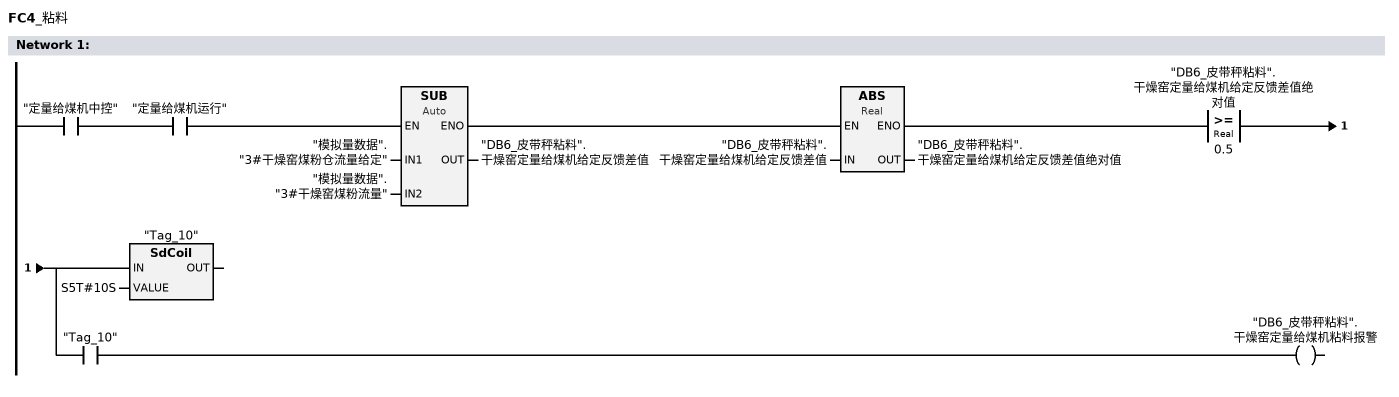
   // no SCL statement known for SdCoil: written as a call
   #_w1 := "定量给煤机中控" AND "定量给煤机运行";
   IF #_w1 THEN
       "DB6_皮带秤粘料".干燥窑定量给煤机给定反馈差值 := "模拟量数据"."3#干燥窑煤粉仓流量给定" - "模拟量数据"."3#干燥窑煤粉流量";
       "DB6_皮带秤粘料".干燥窑定量给煤机给定反馈差值绝对值 := ABS("DB6_皮带秤粘料".干燥窑定量给煤机给定反馈差值);
   END_IF;
   #_w2 := #_w1 AND ("DB6_皮带秤粘料".干燥窑定量给煤机给定反馈差值绝对值 >= 0.5);
   SdCoil(in := #_w2, value := S5T#10S, operand := "Tag_10");
   "DB6_皮带秤粘料".干燥窑定量给煤机粘料报警 := #_w2 AND "Tag_10";
END_REGION
END_FUNCTION

FUNCTION "澳泰温度巡检仪" : Void   // FC5, LAD
{ S7_Optimized_Access := 'FALSE' }
VERSION : 0.1
BEGIN

REGION Network 1
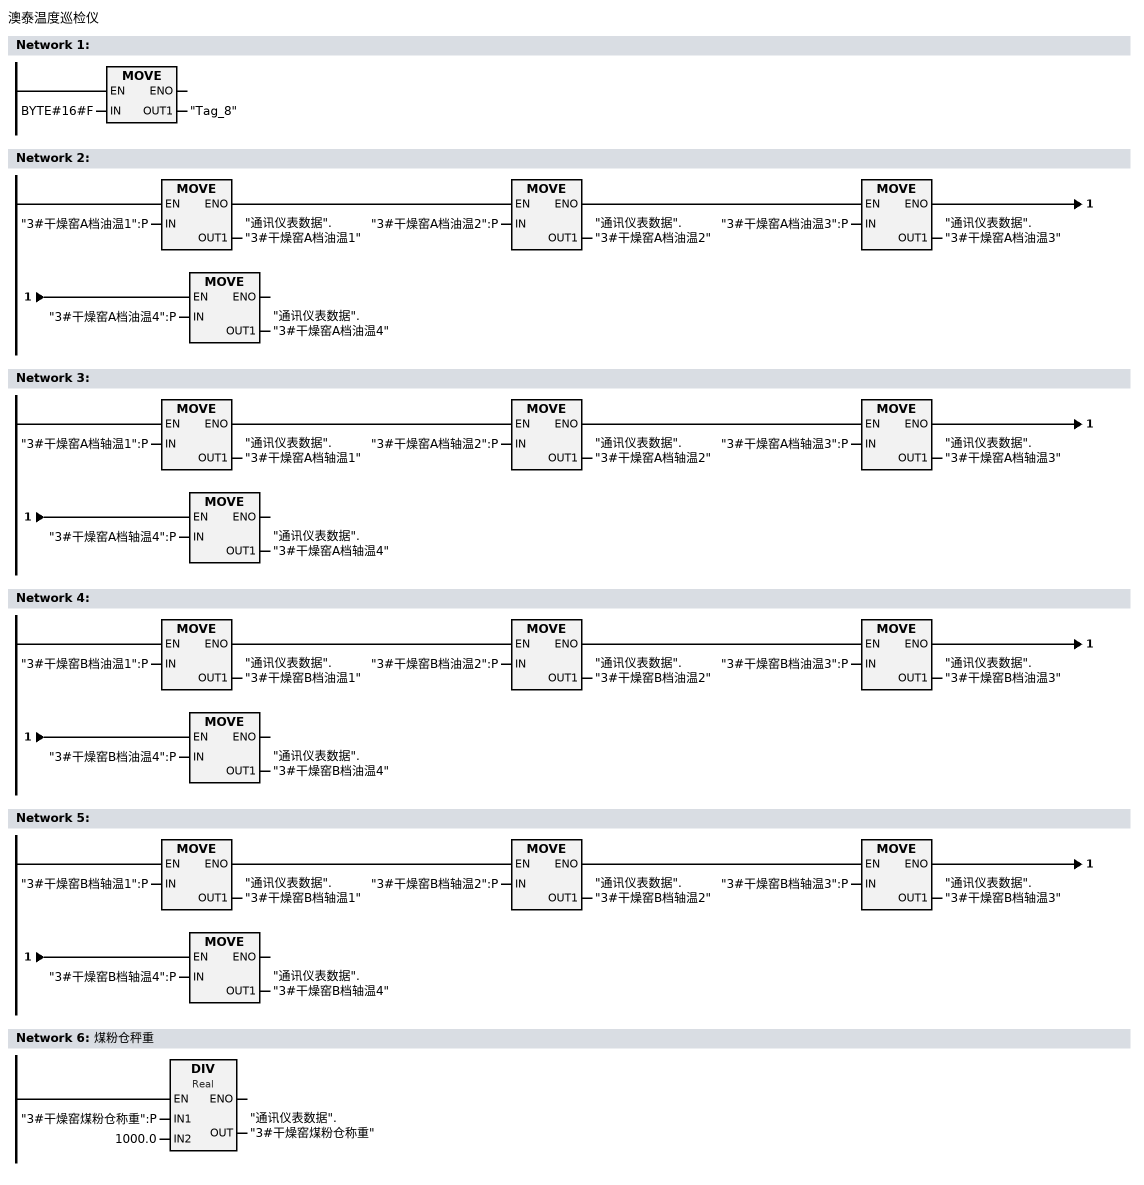
   RUNG wire#powerrail
      { S7_GenerateENO := "TRUE" } Move(in := BYTE#16#F, out1 => "Tag_8")
   END_RUNG
   // the same network as SCL:
   "Tag_8" := BYTE#16#F;
END_REGION

REGION Network 2
   RUNG wire#powerrail
      { S7_GenerateENO := "TRUE" } Move(in := "3#干燥窑A档油温1":P, out1 => "通讯仪表数据"."3#干燥窑A档油温1")
      { S7_GenerateENO := "TRUE" } Move(in := "3#干燥窑A档油温2":P, out1 => "通讯仪表数据"."3#干燥窑A档油温2")
      { S7_GenerateENO := "TRUE" } Move(in := "3#干燥窑A档油温3":P, out1 => "通讯仪表数据"."3#干燥窑A档油温3")
      { S7_GenerateENO := "TRUE" } Move(in := "3#干燥窑A档油温4":P, out1 => "通讯仪表数据"."3#干燥窑A档油温4")
   END_RUNG
   // the same network as SCL:
   // ENO of a box is taken as its EN; it also drops when the box reports an error
   "通讯仪表数据"."3#干燥窑A档油温1" := "3#干燥窑A档油温1":P;
   "通讯仪表数据"."3#干燥窑A档油温2" := "3#干燥窑A档油温2":P;
   "通讯仪表数据"."3#干燥窑A档油温3" := "3#干燥窑A档油温3":P;
   "通讯仪表数据"."3#干燥窑A档油温4" := "3#干燥窑A档油温4":P;
END_REGION

REGION Network 3
   RUNG wire#powerrail
      { S7_GenerateENO := "TRUE" } Move(in := "3#干燥窑A档轴温1":P, out1 => "通讯仪表数据"."3#干燥窑A档轴温1")
      { S7_GenerateENO := "TRUE" } Move(in := "3#干燥窑A档轴温2":P, out1 => "通讯仪表数据"."3#干燥窑A档轴温2")
      { S7_GenerateENO := "TRUE" } Move(in := "3#干燥窑A档轴温3":P, out1 => "通讯仪表数据"."3#干燥窑A档轴温3")
      { S7_GenerateENO := "TRUE" } Move(in := "3#干燥窑A档轴温4":P, out1 => "通讯仪表数据"."3#干燥窑A档轴温4")
   END_RUNG
   // the same network as SCL:
   // ENO of a box is taken as its EN; it also drops when the box reports an error
   "通讯仪表数据"."3#干燥窑A档轴温1" := "3#干燥窑A档轴温1":P;
   "通讯仪表数据"."3#干燥窑A档轴温2" := "3#干燥窑A档轴温2":P;
   "通讯仪表数据"."3#干燥窑A档轴温3" := "3#干燥窑A档轴温3":P;
   "通讯仪表数据"."3#干燥窑A档轴温4" := "3#干燥窑A档轴温4":P;
END_REGION

REGION Network 4
   RUNG wire#powerrail
      { S7_GenerateENO := "TRUE" } Move(in := "3#干燥窑B档油温1":P, out1 => "通讯仪表数据"."3#干燥窑B档油温1")
      { S7_GenerateENO := "TRUE" } Move(in := "3#干燥窑B档油温2":P, out1 => "通讯仪表数据"."3#干燥窑B档油温2")
      { S7_GenerateENO := "TRUE" } Move(in := "3#干燥窑B档油温3":P, out1 => "通讯仪表数据"."3#干燥窑B档油温3")
      { S7_GenerateENO := "TRUE" } Move(in := "3#干燥窑B档油温4":P, out1 => "通讯仪表数据"."3#干燥窑B档油温4")
   END_RUNG
   // the same network as SCL:
   // ENO of a box is taken as its EN; it also drops when the box reports an error
   "通讯仪表数据"."3#干燥窑B档油温1" := "3#干燥窑B档油温1":P;
   "通讯仪表数据"."3#干燥窑B档油温2" := "3#干燥窑B档油温2":P;
   "通讯仪表数据"."3#干燥窑B档油温3" := "3#干燥窑B档油温3":P;
   "通讯仪表数据"."3#干燥窑B档油温4" := "3#干燥窑B档油温4":P;
END_REGION

REGION Network 5
   RUNG wire#powerrail
      { S7_GenerateENO := "TRUE" } Move(in := "3#干燥窑B档轴温1":P, out1 => "通讯仪表数据"."3#干燥窑B档轴温1")
      { S7_GenerateENO := "TRUE" } Move(in := "3#干燥窑B档轴温2":P, out1 => "通讯仪表数据"."3#干燥窑B档轴温2")
      { S7_GenerateENO := "TRUE" } Move(in := "3#干燥窑B档轴温3":P, out1 => "通讯仪表数据"."3#干燥窑B档轴温3")
      { S7_GenerateENO := "TRUE" } Move(in := "3#干燥窑B档轴温4":P, out1 => "通讯仪表数据"."3#干燥窑B档轴温4")
   END_RUNG
   // the same network as SCL:
   // ENO of a box is taken as its EN; it also drops when the box reports an error
   "通讯仪表数据"."3#干燥窑B档轴温1" := "3#干燥窑B档轴温1":P;
   "通讯仪表数据"."3#干燥窑B档轴温2" := "3#干燥窑B档轴温2":P;
   "通讯仪表数据"."3#干燥窑B档轴温3" := "3#干燥窑B档轴温3":P;
   "通讯仪表数据"."3#干燥窑B档轴温4" := "3#干燥窑B档轴温4":P;
END_REGION

REGION Network 6: 煤粉仓秤重
   RUNG wire#powerrail
      { S7_Templates := "SrcType := Real" } Div(in1 := "3#干燥窑煤粉仓称重":P, in2 := 1000.0, out => "通讯仪表数据"."3#干燥窑煤粉仓称重")
   END_RUNG
   // the same network as SCL:
   "通讯仪表数据"."3#干燥窑煤粉仓称重" := "3#干燥窑煤粉仓称重":P / 1000.0;
END_REGION
END_FUNCTION

FUNCTION "3#4#干燥窑皮带联锁信号" : Void   // FC16, LAD
{ S7_Optimized_Access := 'FALSE' }
VERSION : 0.1
BEGIN

REGION Network 1
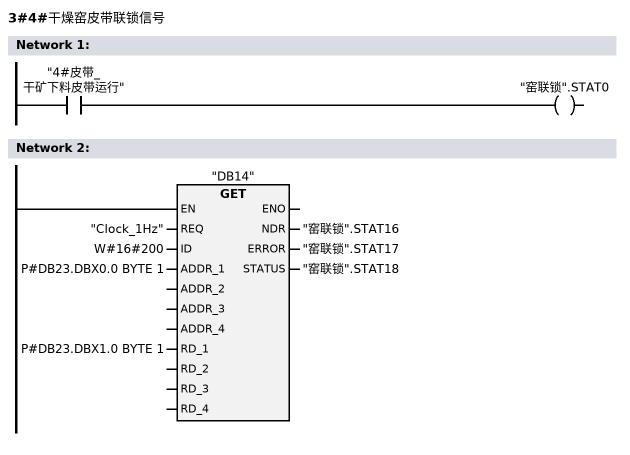
   RUNG wire#powerrail
      Contact( "4#皮带_干矿下料皮带运行" )
      Coil( "窑联锁".STAT0 )
   END_RUNG
   // the same network as SCL:
   "窑联锁".STAT0 := "4#皮带_干矿下料皮带运行";
END_REGION

REGION Network 2
   "DB14"(REQ := "Clock_1Hz",   // GET
          ID := W#16#200,
          ADDR_1 := P#DB23.DBX0.0 BYTE 1,
          RD_1 := P#DB23.DBX1.0 BYTE 1,
          NDR => "窑联锁".STAT16,
          ERROR => "窑联锁".STAT17,
          STATUS => "窑联锁".STAT18);
END_REGION
END_FUNCTION

FUNCTION "模拟量转换" : Void   // FC21, LAD
{ S7_Optimized_Access := 'FALSE' }
VERSION : 0.1
BEGIN

REGION Network 1
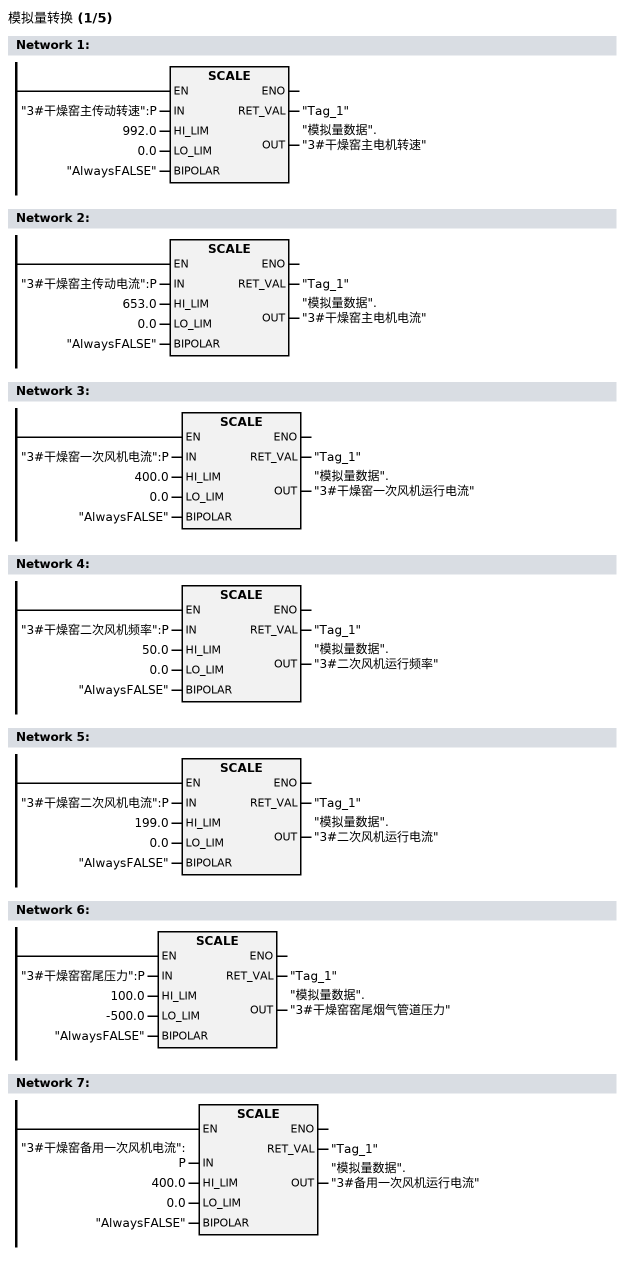
   "Tag_1" := SCALE(IN := "3#干燥窑主传动转速":P,
                    HI_LIM := 992.0,
                    LO_LIM := 0.0,
                    BIPOLAR := "AlwaysFALSE",
                    OUT => "模拟量数据"."3#干燥窑主电机转速");
END_REGION

REGION Network 2
   "Tag_1" := SCALE(IN := "3#干燥窑主传动电流":P,
                    HI_LIM := 653.0,
                    LO_LIM := 0.0,
                    BIPOLAR := "AlwaysFALSE",
                    OUT => "模拟量数据"."3#干燥窑主电机电流");
END_REGION

REGION Network 3
   "Tag_1" := SCALE(IN := "3#干燥窑一次风机电流":P,
                    HI_LIM := 400.0,
                    LO_LIM := 0.0,
                    BIPOLAR := "AlwaysFALSE",
                    OUT => "模拟量数据"."3#干燥窑一次风机运行电流");
END_REGION

REGION Network 4
   "Tag_1" := SCALE(IN := "3#干燥窑二次风机频率":P,
                    HI_LIM := 50.0,
                    LO_LIM := 0.0,
                    BIPOLAR := "AlwaysFALSE",
                    OUT => "模拟量数据"."3#二次风机运行频率");
END_REGION

REGION Network 5
   "Tag_1" := SCALE(IN := "3#干燥窑二次风机电流":P,
                    HI_LIM := 199.0,
                    LO_LIM := 0.0,
                    BIPOLAR := "AlwaysFALSE",
                    OUT => "模拟量数据"."3#二次风机运行电流");
END_REGION

REGION Network 6
   "Tag_1" := SCALE(IN := "3#干燥窑窑尾压力":P,
                    HI_LIM := 100.0,
                    LO_LIM := -500.0,
                    BIPOLAR := "AlwaysFALSE",
                    OUT => "模拟量数据"."3#干燥窑窑尾烟气管道压力");
END_REGION

REGION Network 7
   "Tag_1" := SCALE(IN := "3#干燥窑备用一次风机电流":P,
                    HI_LIM := 400.0,
                    LO_LIM := 0.0,
                    BIPOLAR := "AlwaysFALSE",
                    OUT => "模拟量数据"."3#备用一次风机运行电流");
END_REGION

REGION Network 8
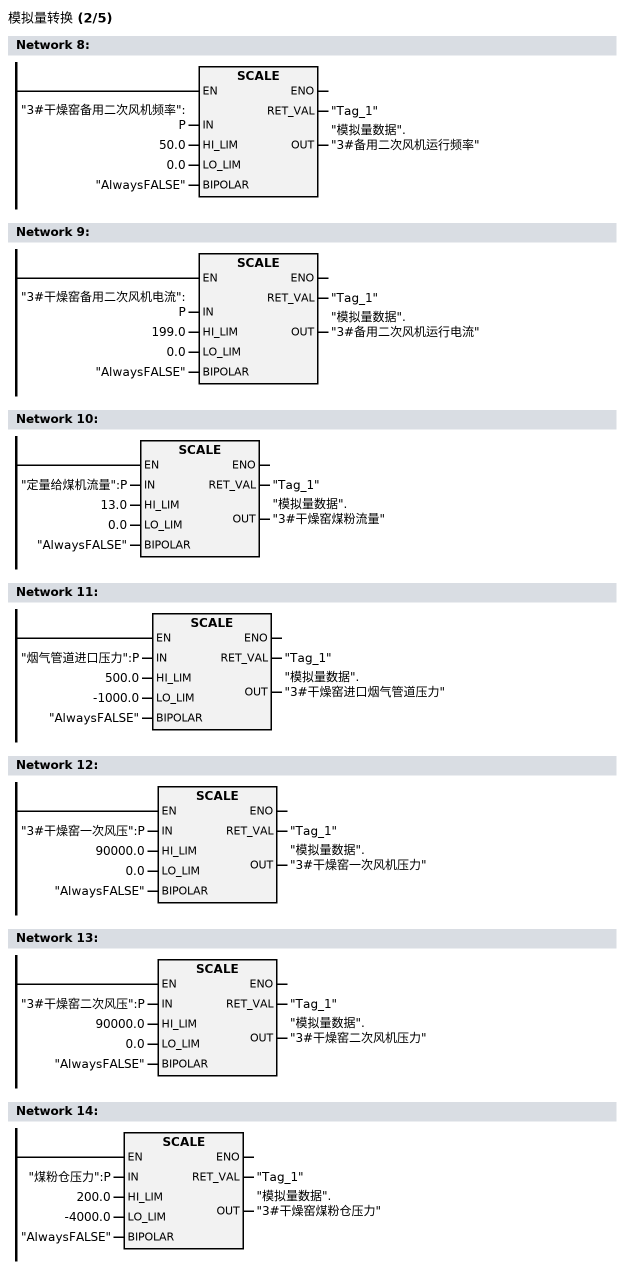
   "Tag_1" := SCALE(IN := "3#干燥窑备用二次风机频率":P,
                    HI_LIM := 50.0,
                    LO_LIM := 0.0,
                    BIPOLAR := "AlwaysFALSE",
                    OUT => "模拟量数据"."3#备用二次风机运行频率");
END_REGION

REGION Network 9
   "Tag_1" := SCALE(IN := "3#干燥窑备用二次风机电流":P,
                    HI_LIM := 199.0,
                    LO_LIM := 0.0,
                    BIPOLAR := "AlwaysFALSE",
                    OUT => "模拟量数据"."3#备用二次风机运行电流");
END_REGION

REGION Network 10
   "Tag_1" := SCALE(IN := "定量给煤机流量":P,
                    HI_LIM := 13.0,
                    LO_LIM := 0.0,
                    BIPOLAR := "AlwaysFALSE",
                    OUT => "模拟量数据"."3#干燥窑煤粉流量");
END_REGION

REGION Network 11
   "Tag_1" := SCALE(IN := "烟气管道进口压力":P,
                    HI_LIM := 500.0,
                    LO_LIM := -1000.0,
                    BIPOLAR := "AlwaysFALSE",
                    OUT => "模拟量数据"."3#干燥窑进口烟气管道压力");
END_REGION

REGION Network 12
   "Tag_1" := SCALE(IN := "3#干燥窑一次风压":P,
                    HI_LIM := 90000.0,
                    LO_LIM := 0.0,
                    BIPOLAR := "AlwaysFALSE",
                    OUT => "模拟量数据"."3#干燥窑一次风机压力");
END_REGION

REGION Network 13
   "Tag_1" := SCALE(IN := "3#干燥窑二次风压":P,
                    HI_LIM := 90000.0,
                    LO_LIM := 0.0,
                    BIPOLAR := "AlwaysFALSE",
                    OUT => "模拟量数据"."3#干燥窑二次风机压力");
END_REGION

REGION Network 14
   "Tag_1" := SCALE(IN := "煤粉仓压力":P,
                    HI_LIM := 200.0,
                    LO_LIM := -4000.0,
                    BIPOLAR := "AlwaysFALSE",
                    OUT => "模拟量数据"."3#干燥窑煤粉仓压力");
END_REGION

REGION Network 15
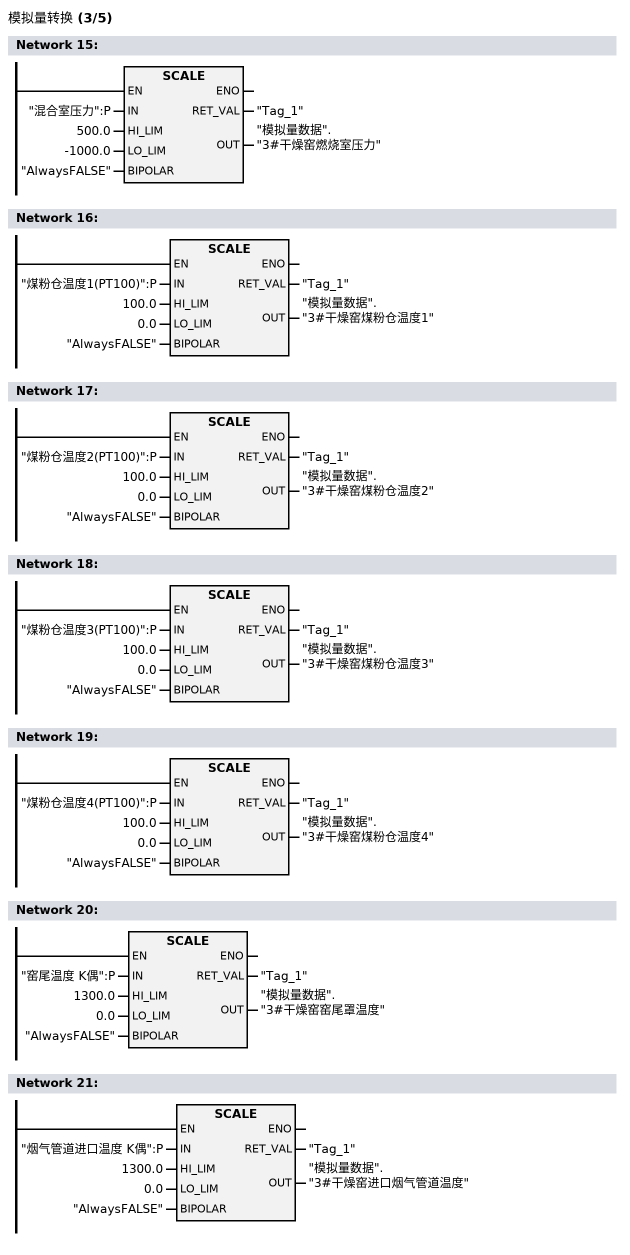
   "Tag_1" := SCALE(IN := "混合室压力":P,
                    HI_LIM := 500.0,
                    LO_LIM := -1000.0,
                    BIPOLAR := "AlwaysFALSE",
                    OUT => "模拟量数据"."3#干燥窑燃烧室压力");
END_REGION

REGION Network 16
   "Tag_1" := SCALE(IN := "煤粉仓温度1(PT100)":P,
                    HI_LIM := 100.0,
                    LO_LIM := 0.0,
                    BIPOLAR := "AlwaysFALSE",
                    OUT => "模拟量数据"."3#干燥窑煤粉仓温度1");
END_REGION

REGION Network 17
   "Tag_1" := SCALE(IN := "煤粉仓温度2(PT100)":P,
                    HI_LIM := 100.0,
                    LO_LIM := 0.0,
                    BIPOLAR := "AlwaysFALSE",
                    OUT => "模拟量数据"."3#干燥窑煤粉仓温度2");
END_REGION

REGION Network 18
   "Tag_1" := SCALE(IN := "煤粉仓温度3(PT100)":P,
                    HI_LIM := 100.0,
                    LO_LIM := 0.0,
                    BIPOLAR := "AlwaysFALSE",
                    OUT => "模拟量数据"."3#干燥窑煤粉仓温度3");
END_REGION

REGION Network 19
   "Tag_1" := SCALE(IN := "煤粉仓温度4(PT100)":P,
                    HI_LIM := 100.0,
                    LO_LIM := 0.0,
                    BIPOLAR := "AlwaysFALSE",
                    OUT => "模拟量数据"."3#干燥窑煤粉仓温度4");
END_REGION

REGION Network 20
   "Tag_1" := SCALE(IN := "窑尾温度 K偶":P,
                    HI_LIM := 1300.0,
                    LO_LIM := 0.0,
                    BIPOLAR := "AlwaysFALSE",
                    OUT => "模拟量数据"."3#干燥窑窑尾罩温度");
END_REGION

REGION Network 21
   "Tag_1" := SCALE(IN := "烟气管道进口温度 K偶":P,
                    HI_LIM := 1300.0,
                    LO_LIM := 0.0,
                    BIPOLAR := "AlwaysFALSE",
                    OUT => "模拟量数据"."3#干燥窑进口烟气管道温度");
END_REGION

REGION Network 22
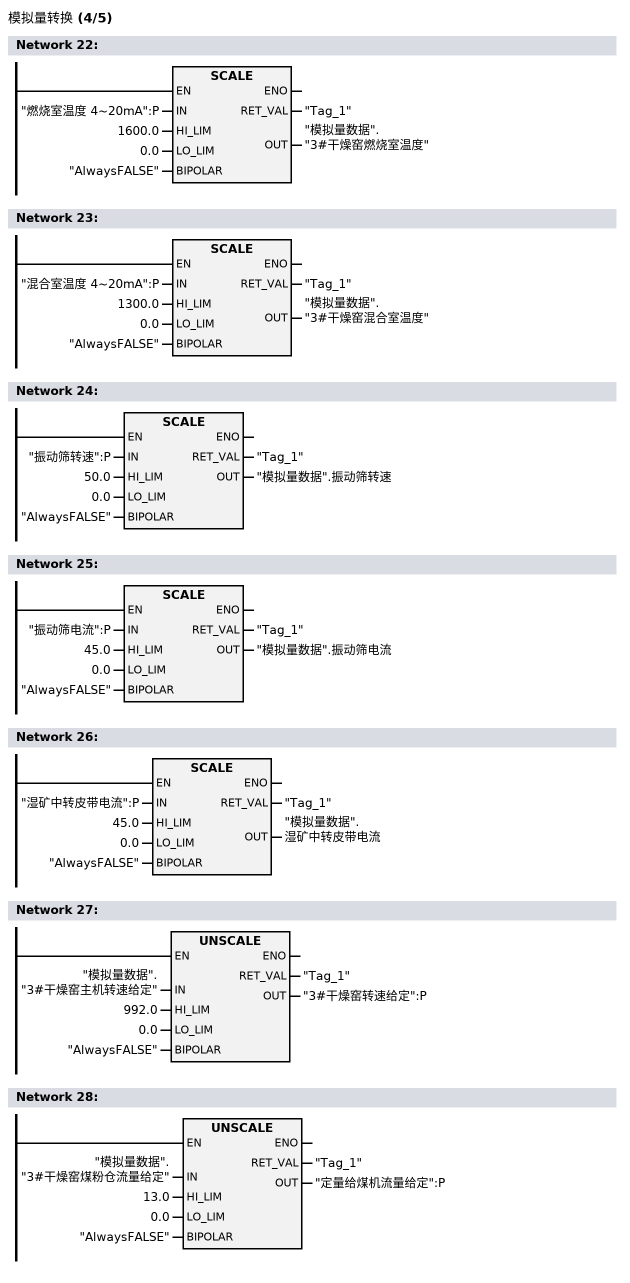
   "Tag_1" := SCALE(IN := "燃烧室温度 4~20mA":P,
                    HI_LIM := 1600.0,
                    LO_LIM := 0.0,
                    BIPOLAR := "AlwaysFALSE",
                    OUT => "模拟量数据"."3#干燥窑燃烧室温度");
END_REGION

REGION Network 23
   "Tag_1" := SCALE(IN := "混合室温度 4~20mA":P,
                    HI_LIM := 1300.0,
                    LO_LIM := 0.0,
                    BIPOLAR := "AlwaysFALSE",
                    OUT => "模拟量数据"."3#干燥窑混合室温度");
END_REGION

REGION Network 24
   "Tag_1" := SCALE(IN := "振动筛转速":P,
                    HI_LIM := 50.0,
                    LO_LIM := 0.0,
                    BIPOLAR := "AlwaysFALSE",
                    OUT => "模拟量数据".振动筛转速);
END_REGION

REGION Network 25
   "Tag_1" := SCALE(IN := "振动筛电流":P,
                    HI_LIM := 45.0,
                    LO_LIM := 0.0,
                    BIPOLAR := "AlwaysFALSE",
                    OUT => "模拟量数据".振动筛电流);
END_REGION

REGION Network 26
   "Tag_1" := SCALE(IN := "湿矿中转皮带电流":P,
                    HI_LIM := 45.0,
                    LO_LIM := 0.0,
                    BIPOLAR := "AlwaysFALSE",
                    OUT => "模拟量数据".湿矿中转皮带电流);
END_REGION

REGION Network 27
   "Tag_1" := UNSCALE(IN := "模拟量数据"."3#干燥窑主机转速给定",
                      HI_LIM := 992.0,
                      LO_LIM := 0.0,
                      BIPOLAR := "AlwaysFALSE",
                      OUT => "3#干燥窑转速给定":P);
END_REGION

REGION Network 28
   "Tag_1" := UNSCALE(IN := "模拟量数据"."3#干燥窑煤粉仓流量给定",
                      HI_LIM := 13.0,
                      LO_LIM := 0.0,
                      BIPOLAR := "AlwaysFALSE",
                      OUT => "定量给煤机流量给定":P);
END_REGION

REGION Network 29
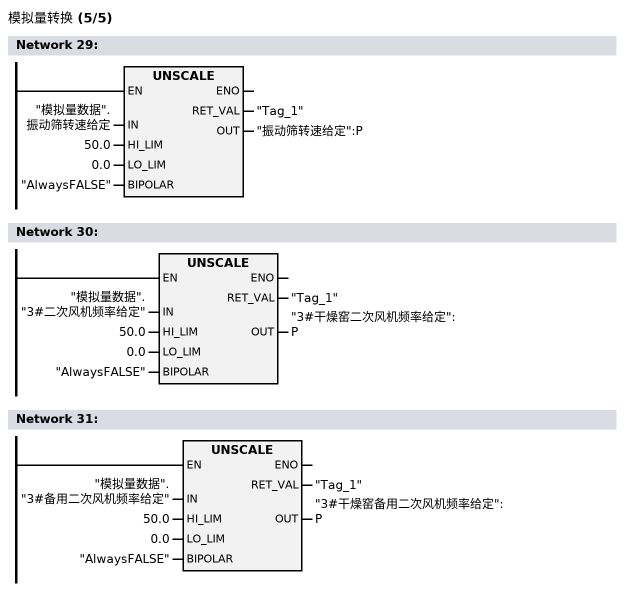
   "Tag_1" := UNSCALE(IN := "模拟量数据".振动筛转速给定,
                      HI_LIM := 50.0,
                      LO_LIM := 0.0,
                      BIPOLAR := "AlwaysFALSE",
                      OUT => "振动筛转速给定":P);
END_REGION

REGION Network 30
   "Tag_1" := UNSCALE(IN := "模拟量数据"."3#二次风机频率给定",
                      HI_LIM := 50.0,
                      LO_LIM := 0.0,
                      BIPOLAR := "AlwaysFALSE",
                      OUT => "3#干燥窑二次风机频率给定":P);
END_REGION

REGION Network 31
   "Tag_1" := UNSCALE(IN := "模拟量数据"."3#备用二次风机频率给定",
                      HI_LIM := 50.0,
                      LO_LIM := 0.0,
                      BIPOLAR := "AlwaysFALSE",
                      OUT => "3#干燥窑备用二次风机频率给定":P);
END_REGION
END_FUNCTION

FUNCTION "皮带机" : Void   // FC22, LAD
{ S7_Optimized_Access := 'FALSE' }
VERSION : 0.1
BEGIN

REGION Network 1
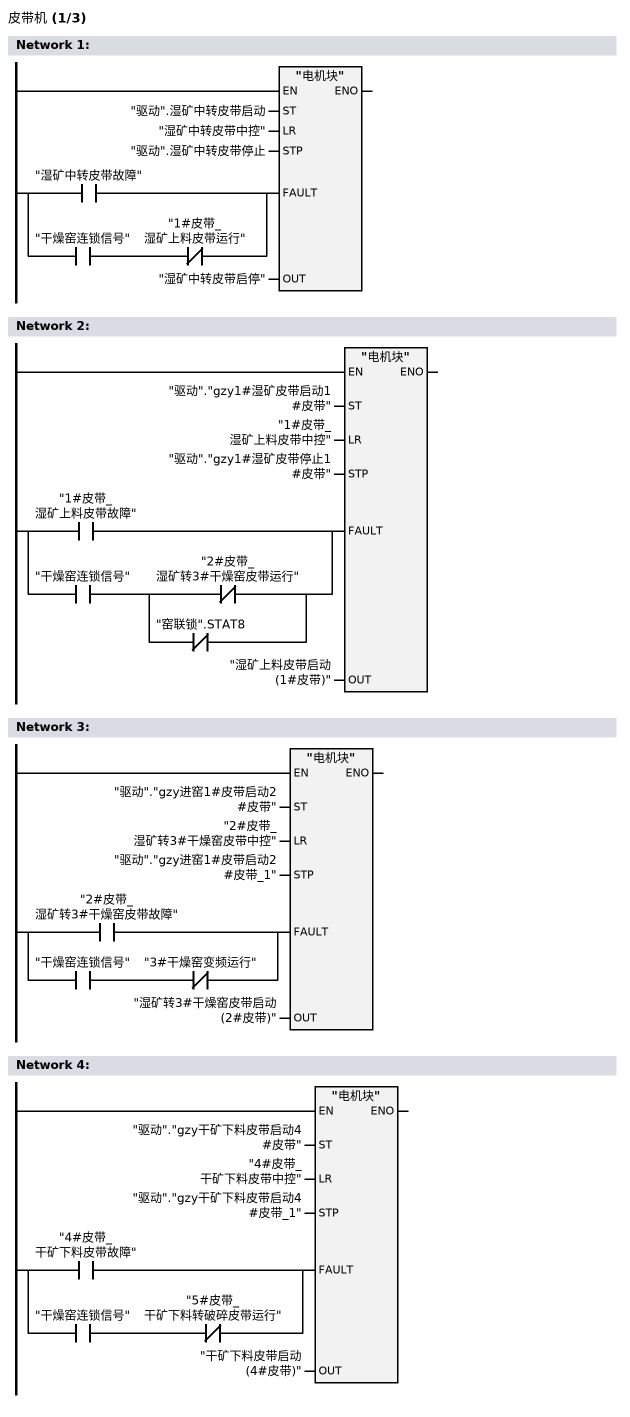
   RUNG wire#powerrail
      "电机块"(FAULT := wire#w1, ST := "驱动".湿矿中转皮带启动, LR := "湿矿中转皮带中控", STP := "驱动".湿矿中转皮带停止, OUT := "湿矿中转皮带启停")
   END_RUNG
   RUNG wire#powerrail
      Contact( "湿矿中转皮带故障" )
   END_RUNG wire#w1
   RUNG wire#powerrail
      Contact( "干燥窑连锁信号" )
      I_Contact( "1#皮带_湿矿上料皮带运行" )
   END_RUNG wire#w1
   // the same network as SCL:
   "电机块"(ST := "驱动".湿矿中转皮带启动,
         LR := "湿矿中转皮带中控",
         STP := "驱动".湿矿中转皮带停止,
         FAULT := "湿矿中转皮带故障" OR ("干燥窑连锁信号" AND NOT "1#皮带_湿矿上料皮带运行"),
         OUT := "湿矿中转皮带启停");
END_REGION

REGION Network 2
   RUNG wire#powerrail
      "电机块"(FAULT := wire#w2, ST := "驱动"."gzy1#湿矿皮带启动1#皮带", LR := "1#皮带_湿矿上料皮带中控", STP := "驱动"."gzy1#湿矿皮带停止1#皮带", OUT := "湿矿上料皮带启动  (1#皮带)")
   END_RUNG
   RUNG wire#powerrail
      Contact( "1#皮带_湿矿上料皮带故障" )
   END_RUNG wire#w2
   RUNG wire#powerrail
      Contact( "干燥窑连锁信号" )
      wire#w1
      I_Contact( "2#皮带_湿矿转3#干燥窑皮带运行" )
   END_RUNG wire#w2
   RUNG wire#w1
      I_Contact( "窑联锁".STAT8 )
   END_RUNG wire#w2
   // the same network as SCL:
   "电机块"(ST := "驱动"."gzy1#湿矿皮带启动1#皮带",
         LR := "1#皮带_湿矿上料皮带中控",
         STP := "驱动"."gzy1#湿矿皮带停止1#皮带",
         FAULT := "1#皮带_湿矿上料皮带故障" OR ("干燥窑连锁信号" AND (NOT "2#皮带_湿矿转3#干燥窑皮带运行" OR NOT "窑联锁".STAT8)),
         OUT := "湿矿上料皮带启动  (1#皮带)");
END_REGION

REGION Network 3
   RUNG wire#powerrail
      "电机块"(FAULT := wire#w1, ST := "驱动"."gzy进窑1#皮带启动2#皮带", LR := "2#皮带_湿矿转3#干燥窑皮带中控", STP := "驱动"."gzy进窑1#皮带启动2#皮带_1", OUT := "湿矿转3#干燥窑皮带启动  (2#皮带)")
   END_RUNG
   RUNG wire#powerrail
      Contact( "2#皮带_湿矿转3#干燥窑皮带故障" )
   END_RUNG wire#w1
   RUNG wire#powerrail
      Contact( "干燥窑连锁信号" )
      I_Contact( "3#干燥窑变频运行" )
   END_RUNG wire#w1
   // the same network as SCL:
   "电机块"(ST := "驱动"."gzy进窑1#皮带启动2#皮带",
         LR := "2#皮带_湿矿转3#干燥窑皮带中控",
         STP := "驱动"."gzy进窑1#皮带启动2#皮带_1",
         FAULT := "2#皮带_湿矿转3#干燥窑皮带故障" OR ("干燥窑连锁信号" AND NOT "3#干燥窑变频运行"),
         OUT := "湿矿转3#干燥窑皮带启动  (2#皮带)");
END_REGION

REGION Network 4
   RUNG wire#powerrail
      "电机块"(FAULT := wire#w1, ST := "驱动"."gzy干矿下料皮带启动4#皮带", LR := "4#皮带_干矿下料皮带中控", STP := "驱动"."gzy干矿下料皮带启动4#皮带_1", OUT := "干矿下料皮带启动  (4#皮带)")
   END_RUNG
   RUNG wire#powerrail
      Contact( "4#皮带_干矿下料皮带故障" )
   END_RUNG wire#w1
   RUNG wire#powerrail
      Contact( "干燥窑连锁信号" )
      I_Contact( "5#皮带_干矿下料转破碎皮带运行" )
   END_RUNG wire#w1
   // the same network as SCL:
   "电机块"(ST := "驱动"."gzy干矿下料皮带启动4#皮带",
         LR := "4#皮带_干矿下料皮带中控",
         STP := "驱动"."gzy干矿下料皮带启动4#皮带_1",
         FAULT := "4#皮带_干矿下料皮带故障" OR ("干燥窑连锁信号" AND NOT "5#皮带_干矿下料转破碎皮带运行"),
         OUT := "干矿下料皮带启动  (4#皮带)");
END_REGION

REGION Network 5
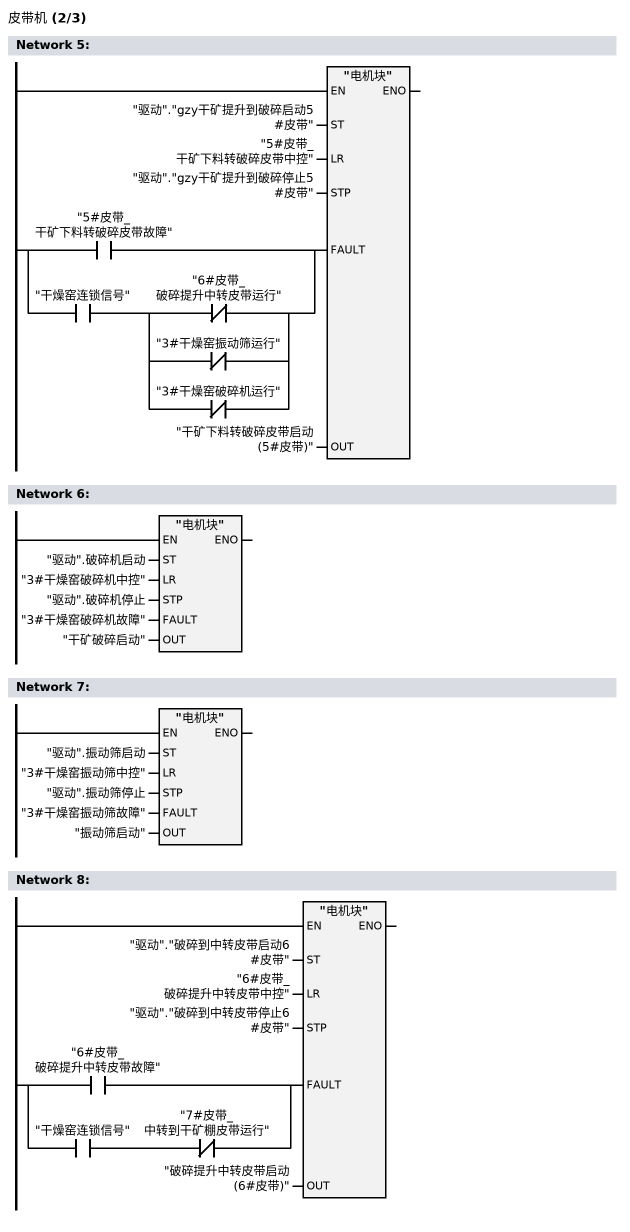
   RUNG wire#powerrail
      "电机块"(FAULT := wire#w2, ST := "驱动"."gzy干矿提升到破碎启动5#皮带", LR := "5#皮带_干矿下料转破碎皮带中控", STP := "驱动"."gzy干矿提升到破碎停止5#皮带", OUT := "干矿下料转破碎皮带启动  (5#皮带)")
   END_RUNG
   RUNG wire#powerrail
      Contact( "5#皮带_干矿下料转破碎皮带故障" )
   END_RUNG wire#w2
   RUNG wire#powerrail
      Contact( "干燥窑连锁信号" )
      wire#w1
      I_Contact( "6#皮带_破碎提升中转皮带运行" )
   END_RUNG wire#w2
   RUNG wire#w1
      I_Contact( "3#干燥窑振动筛运行" )
   END_RUNG wire#w2
   RUNG wire#w1
      I_Contact( "3#干燥窑破碎机运行" )
   END_RUNG wire#w2
   // the same network as SCL:
   "电机块"(ST := "驱动"."gzy干矿提升到破碎启动5#皮带",
         LR := "5#皮带_干矿下料转破碎皮带中控",
         STP := "驱动"."gzy干矿提升到破碎停止5#皮带",
         FAULT := "5#皮带_干矿下料转破碎皮带故障" OR ("干燥窑连锁信号" AND (NOT "6#皮带_破碎提升中转皮带运行" OR NOT "3#干燥窑振动筛运行" OR NOT "3#干燥窑破碎机运行")),
         OUT := "干矿下料转破碎皮带启动  (5#皮带)");
END_REGION

REGION Network 6
   RUNG wire#powerrail
      "电机块"(ST := "驱动".破碎机启动, LR := "3#干燥窑破碎机中控", STP := "驱动".破碎机停止, FAULT := "3#干燥窑破碎机故障", OUT := "干矿破碎启动")
   END_RUNG
   // the same network as SCL:
   "电机块"(ST := "驱动".破碎机启动, LR := "3#干燥窑破碎机中控", STP := "驱动".破碎机停止, FAULT := "3#干燥窑破碎机故障", OUT := "干矿破碎启动");
END_REGION

REGION Network 7
   RUNG wire#powerrail
      "电机块"(ST := "驱动".振动筛启动, LR := "3#干燥窑振动筛中控", STP := "驱动".振动筛停止, FAULT := "3#干燥窑振动筛故障", OUT := "振动筛启动")
   END_RUNG
   // the same network as SCL:
   "电机块"(ST := "驱动".振动筛启动, LR := "3#干燥窑振动筛中控", STP := "驱动".振动筛停止, FAULT := "3#干燥窑振动筛故障", OUT := "振动筛启动");
END_REGION

REGION Network 8
   RUNG wire#powerrail
      "电机块"(FAULT := wire#w1, ST := "驱动"."破碎到中转皮带启动6#皮带", LR := "6#皮带_破碎提升中转皮带中控", STP := "驱动"."破碎到中转皮带停止6#皮带", OUT := "破碎提升中转皮带启动  (6#皮带)")
   END_RUNG
   RUNG wire#powerrail
      Contact( "6#皮带_破碎提升中转皮带故障" )
   END_RUNG wire#w1
   RUNG wire#powerrail
      Contact( "干燥窑连锁信号" )
      I_Contact( "7#皮带_中转到干矿棚皮带运行" )
   END_RUNG wire#w1
   // the same network as SCL:
   "电机块"(ST := "驱动"."破碎到中转皮带启动6#皮带",
         LR := "6#皮带_破碎提升中转皮带中控",
         STP := "驱动"."破碎到中转皮带停止6#皮带",
         FAULT := "6#皮带_破碎提升中转皮带故障" OR ("干燥窑连锁信号" AND NOT "7#皮带_中转到干矿棚皮带运行"),
         OUT := "破碎提升中转皮带启动  (6#皮带)");
END_REGION

REGION Network 9
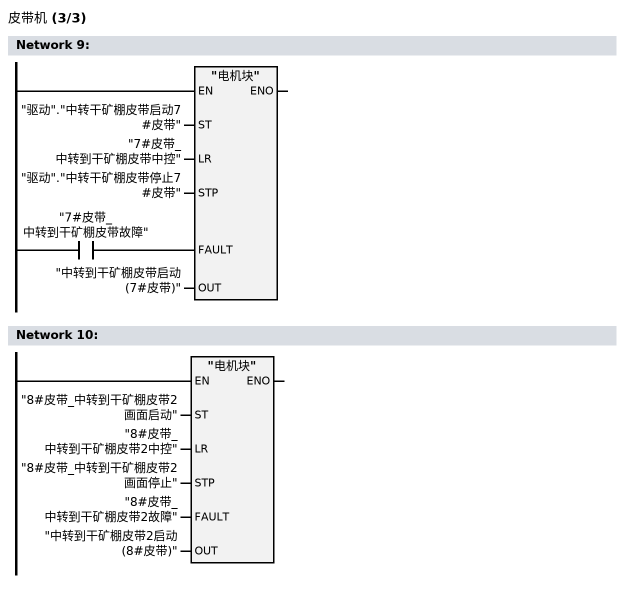
   RUNG wire#powerrail
      "电机块"(FAULT := wire#w1, ST := "驱动"."中转干矿棚皮带启动7#皮带", LR := "7#皮带_中转到干矿棚皮带中控", STP := "驱动"."中转干矿棚皮带停止7#皮带", OUT := "中转到干矿棚皮带启动  (7#皮带)")
   END_RUNG
   RUNG wire#powerrail
      Contact( "7#皮带_中转到干矿棚皮带故障" )
   END_RUNG wire#w1
   // the same network as SCL:
   "电机块"(ST := "驱动"."中转干矿棚皮带启动7#皮带",
         LR := "7#皮带_中转到干矿棚皮带中控",
         STP := "驱动"."中转干矿棚皮带停止7#皮带",
         FAULT := "7#皮带_中转到干矿棚皮带故障",
         OUT := "中转到干矿棚皮带启动  (7#皮带)");
END_REGION

REGION Network 10
   RUNG wire#powerrail
      "电机块"(ST := "8#皮带_中转到干矿棚皮带2画面启动", LR := "8#皮带_中转到干矿棚皮带2中控", STP := "8#皮带_中转到干矿棚皮带2画面停止", FAULT := "8#皮带_中转到干矿棚皮带2故障", OUT := "中转到干矿棚皮带2启动  (8#皮带)")
   END_RUNG
   // the same network as SCL:
   "电机块"(ST := "8#皮带_中转到干矿棚皮带2画面启动",
         LR := "8#皮带_中转到干矿棚皮带2中控",
         STP := "8#皮带_中转到干矿棚皮带2画面停止",
         FAULT := "8#皮带_中转到干矿棚皮带2故障",
         OUT := "中转到干矿棚皮带2启动  (8#皮带)");
END_REGION
END_FUNCTION

FUNCTION "给煤机累计" : Void   // FC23, LAD
{ S7_Optimized_Access := 'FALSE' }
VERSION : 0.1
   VAR_TEMP   // added for the SCL form of the ladder/FBD networks
      _w1 : Bool;
      _w2 : Bool;
   END_VAR
BEGIN

REGION Network 1
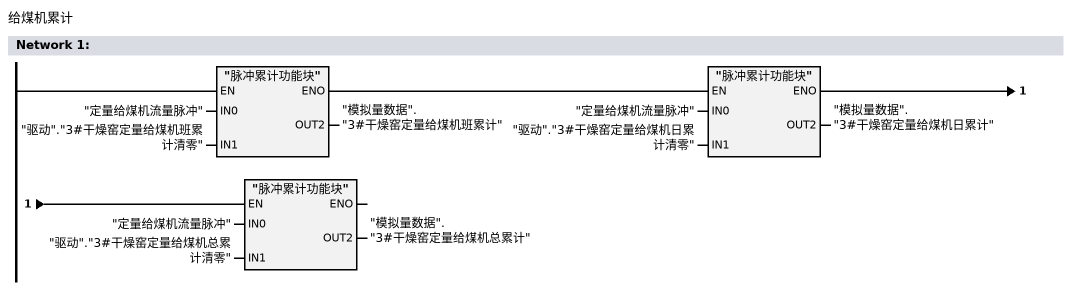
   RUNG wire#powerrail
      "脉冲累计功能块"(IN0 := "定量给煤机流量脉冲", IN1 := "驱动"."3#干燥窑定量给煤机班累计清零", OUT2 => "模拟量数据"."3#干燥窑定量给煤机班累计")
      "脉冲累计功能块"(IN0 := "定量给煤机流量脉冲", IN1 := "驱动"."3#干燥窑定量给煤机日累计清零", OUT2 => "模拟量数据"."3#干燥窑定量给煤机日累计")
      "脉冲累计功能块"(IN0 := "定量给煤机流量脉冲", IN1 := "驱动"."3#干燥窑定量给煤机总累计清零", OUT2 => "模拟量数据"."3#干燥窑定量给煤机总累计")
   END_RUNG
   // the same network as SCL:
   "脉冲累计功能块"(IN0 := "定量给煤机流量脉冲", IN1 := "驱动"."3#干燥窑定量给煤机班累计清零", OUT2 => "模拟量数据"."3#干燥窑定量给煤机班累计", ENO => #_w1);
   "脉冲累计功能块"(EN := #_w1,
             IN0 := "定量给煤机流量脉冲",
             IN1 := "驱动"."3#干燥窑定量给煤机日累计清零",
             OUT2 => "模拟量数据"."3#干燥窑定量给煤机日累计",
             ENO => #_w2);
   IF #_w2 THEN
       "脉冲累计功能块"(IN0 := "定量给煤机流量脉冲", IN1 := "驱动"."3#干燥窑定量给煤机总累计清零", OUT2 => "模拟量数据"."3#干燥窑定量给煤机总累计");
   END_IF;
END_REGION
END_FUNCTION

FUNCTION "FC40_DATA_ALARM" : Void   // FC40, LAD
{ S7_Optimized_Access := 'TRUE' }
VERSION : 0.1
BEGIN

REGION Network 1
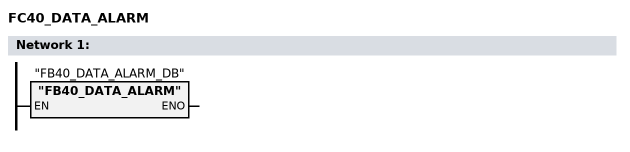
   RUNG wire#powerrail
      "FB40_DATA_ALARM_DB"()
   END_RUNG
   // the same network as SCL:
   "FB40_DATA_ALARM_DB"();   // "FB40_DATA_ALARM"
END_REGION
END_FUNCTION

FUNCTION "脉冲累计功能块" : Void   // FC116, LAD
{ S7_Optimized_Access := 'FALSE' }
VERSION : 0.1
   VAR_INPUT
      IN0 : Bool;
      IN1 : Bool;
   END_VAR
   VAR_OUTPUT
      OUT2 : Real;
   END_VAR
   VAR_TEMP
      TEMP3 : Bool;
      TEMP4 : Real;
      TEMP5 : Real;
      TEMP6 : Real;
   END_VAR
   VAR_TEMP   // added for the SCL form of the ladder/FBD networks
      _w1 : Bool;
   END_VAR
BEGIN

REGION Network 2
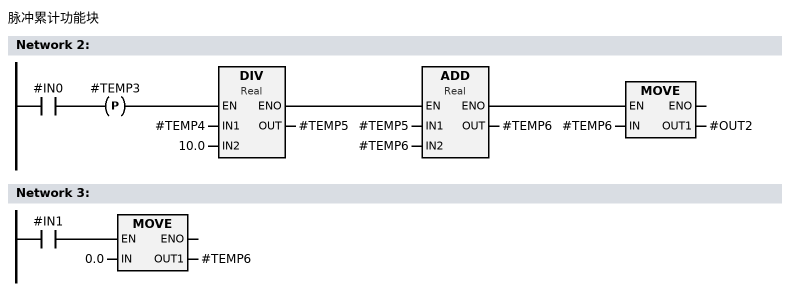
   RUNG wire#powerrail
      Contact( #IN0 )
      P_Trig( #TEMP3 )
      { S7_Templates := "SrcType := Real"; S7_GenerateENO := "TRUE" } Div(in1 := #TEMP4, in2 := 10.0, out => #TEMP5)
      { S7_Templates := "SrcType := Real"; S7_GenerateENO := "TRUE" } Add(in1 := #TEMP5, in2 := #TEMP6, out => #TEMP6)
      { S7_GenerateENO := "TRUE" } Move(in := #TEMP6, out1 => #OUT2)
   END_RUNG
   // the same network as SCL:
   // ENO of a box is taken as its EN; it also drops when the box reports an error
   #_w1 := #IN0 AND NOT #TEMP3;   // rising edge
   #TEMP3 := #IN0;
   IF #_w1 THEN
       #TEMP5 := #TEMP4 / 10.0;
       #TEMP6 := #TEMP5 + #TEMP6;
       #OUT2 := #TEMP6;
   END_IF;
END_REGION

REGION Network 3
   RUNG wire#powerrail
      Contact( #IN1 )
      { S7_GenerateENO := "TRUE" } Move(in := 0.0, out1 => #TEMP6)
   END_RUNG
   // the same network as SCL:
   IF #IN1 THEN #TEMP6 := 0.0; END_IF;
END_REGION

REGION Network 4 (STL)
         SET;
         SAVE;
END_REGION
END_FUNCTION

ORGANIZATION_BLOCK "Main"   // OB1, LAD, ProgramCycle
TITLE = "Main Program Sweep (Cycle)"
{ S7_Optimized_Access := 'TRUE' }
VERSION : 0.1
   VAR_INPUT
      Initial_Call : Bool;   // Initial call of this OB
      Remanence : Bool;   // =True, if remanent data are available
   END_VAR
BEGIN

REGION Network 1
